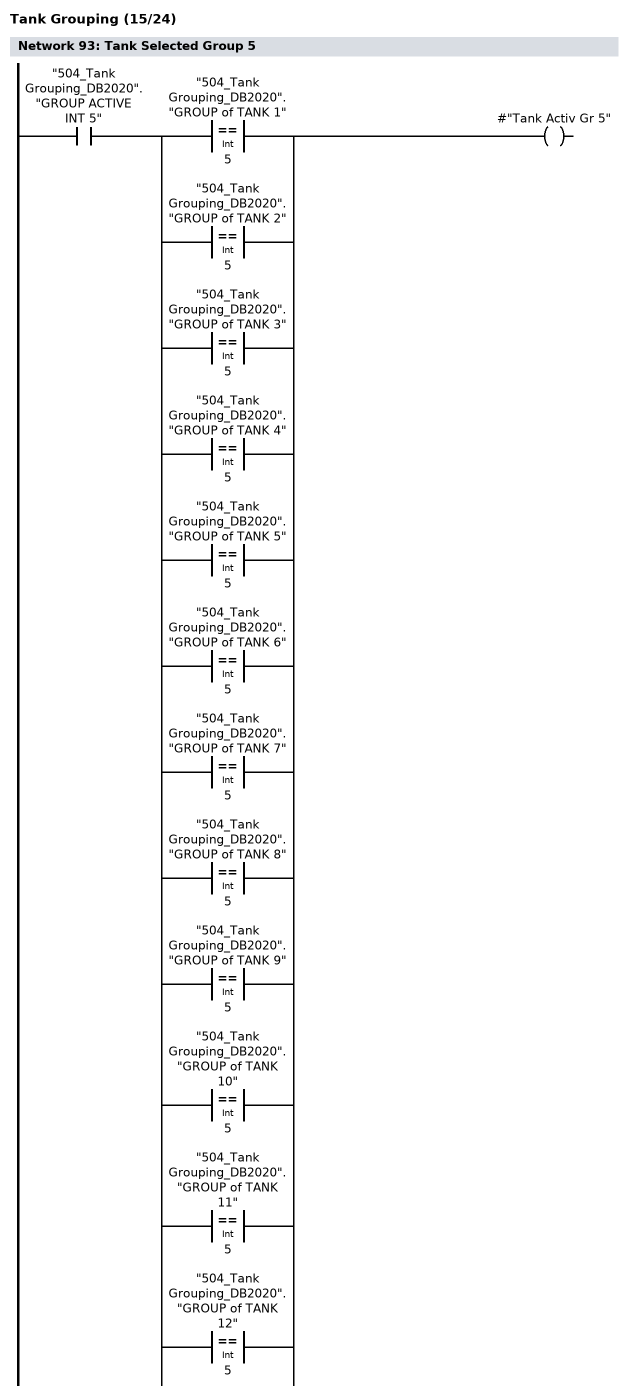
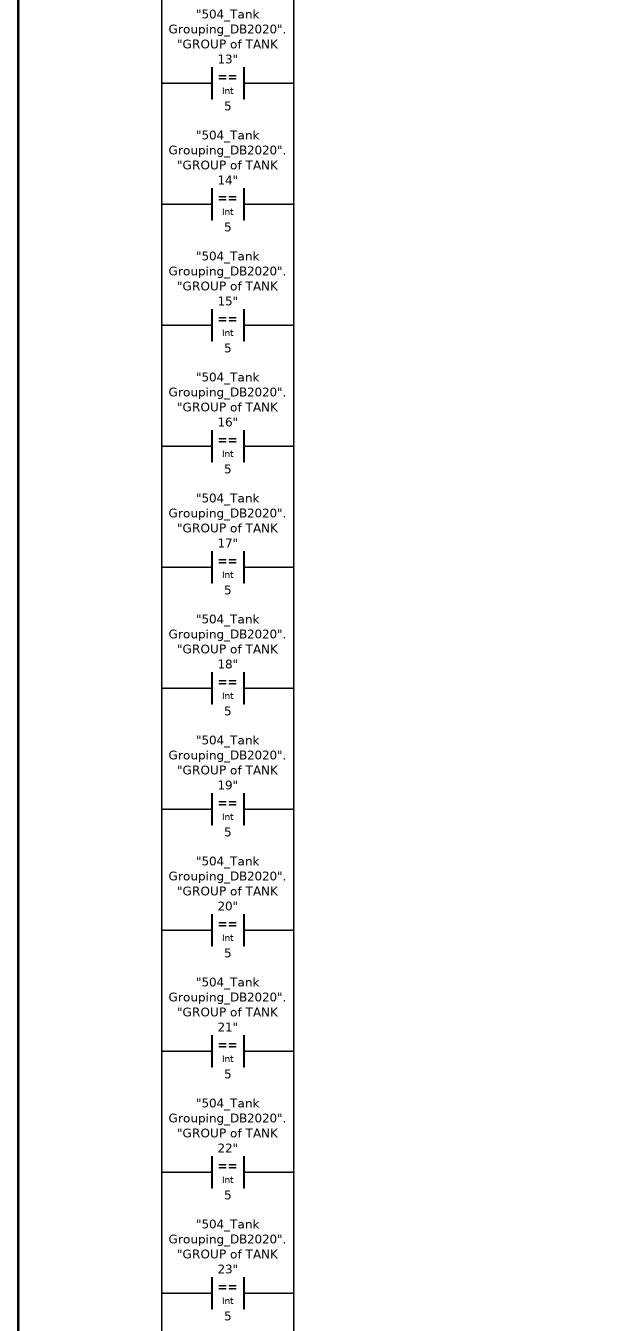
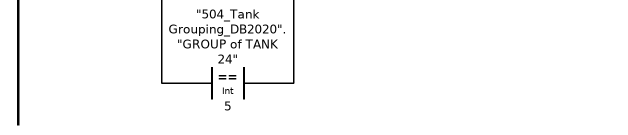
   RUNG wire#powerrail
      Contact( "504_Tank Grouping_DB2020"."GROUP ACTIVE INT 5" )
      wire#w1
      { S7_Templates := "SrcType := Int" } EQ_Contact(in1 := "504_Tank Grouping_DB2020"."GROUP of TANK 1", in2 := 5)
      wire#w2
      Coil( #"Tank Activ Gr 5" )
   END_RUNG
   RUNG wire#w1
      { S7_Templates := "SrcType := Int" } EQ_Contact(in1 := "504_Tank Grouping_DB2020"."GROUP of TANK 2", in2 := 5)
   END_RUNG wire#w2
   RUNG wire#w1
      { S7_Templates := "SrcType := Int" } EQ_Contact(in1 := "504_Tank Grouping_DB2020"."GROUP of TANK 3", in2 := 5)
   END_RUNG wire#w2
   RUNG wire#w1
      { S7_Templates := "SrcType := Int" } EQ_Contact(in1 := "504_Tank Grouping_DB2020"."GROUP of TANK 4", in2 := 5)
   END_RUNG wire#w2
   RUNG wire#w1
      { S7_Templates := "SrcType := Int" } EQ_Contact(in1 := "504_Tank Grouping_DB2020"."GROUP of TANK 5", in2 := 5)
   END_RUNG wire#w2
   RUNG wire#w1
      { S7_Templates := "SrcType := Int" } EQ_Contact(in1 := "504_Tank Grouping_DB2020"."GROUP of TANK 6", in2 := 5)
   END_RUNG wire#w2
   RUNG wire#w1
      { S7_Templates := "SrcType := Int" } EQ_Contact(in1 := "504_Tank Grouping_DB2020"."GROUP of TANK 7", in2 := 5)
   END_RUNG wire#w2
   RUNG wire#w1
      { S7_Templates := "SrcType := Int" } EQ_Contact(in1 := "504_Tank Grouping_DB2020"."GROUP of TANK 8", in2 := 5)
   END_RUNG wire#w2
   RUNG wire#w1
      { S7_Templates := "SrcType := Int" } EQ_Contact(in1 := "504_Tank Grouping_DB2020"."GROUP of TANK 9", in2 := 5)
   END_RUNG wire#w2
   RUNG wire#w1
      { S7_Templates := "SrcType := Int" } EQ_Contact(in1 := "504_Tank Grouping_DB2020"."GROUP of TANK 10", in2 := 5)
   END_RUNG wire#w2
   RUNG wire#w1
      { S7_Templates := "SrcType := Int" } EQ_Contact(in1 := "504_Tank Grouping_DB2020"."GROUP of TANK 11", in2 := 5)
   END_RUNG wire#w2
   RUNG wire#w1
      { S7_Templates := "SrcType := Int" } EQ_Contact(in1 := "504_Tank Grouping_DB2020"."GROUP of TANK 12", in2 := 5)
   END_RUNG wire#w2
   RUNG wire#w1
      { S7_Templates := "SrcType := Int" } EQ_Contact(in1 := "504_Tank Grouping_DB2020"."GROUP of TANK 13", in2 := 5)
   END_RUNG wire#w2
   RUNG wire#w1
      { S7_Templates := "SrcType := Int" } EQ_Contact(in1 := "504_Tank Grouping_DB2020"."GROUP of TANK 14", in2 := 5)
   END_RUNG wire#w2
   RUNG wire#w1
      { S7_Templates := "SrcType := Int" } EQ_Contact(in1 := "504_Tank Grouping_DB2020"."GROUP of TANK 15", in2 := 5)
   END_RUNG wire#w2
   RUNG wire#w1
      { S7_Templates := "SrcType := Int" } EQ_Contact(in1 := "504_Tank Grouping_DB2020"."GROUP of TANK 16", in2 := 5)
   END_RUNG wire#w2
   RUNG wire#w1
      { S7_Templates := "SrcType := Int" } EQ_Contact(in1 := "504_Tank Grouping_DB2020"."GROUP of TANK 17", in2 := 5)
   END_RUNG wire#w2
   RUNG wire#w1
      { S7_Templates := "SrcType := Int" } EQ_Contact(in1 := "504_Tank Grouping_DB2020"."GROUP of TANK 18", in2 := 5)
   END_RUNG wire#w2
   RUNG wire#w1
      { S7_Templates := "SrcType := Int" } EQ_Contact(in1 := "504_Tank Grouping_DB2020"."GROUP of TANK 19", in2 := 5)
   END_RUNG wire#w2
   RUNG wire#w1
      { S7_Templates := "SrcType := Int" } EQ_Contact(in1 := "504_Tank Grouping_DB2020"."GROUP of TANK 20", in2 := 5)
   END_RUNG wire#w2
   RUNG wire#w1
      { S7_Templates := "SrcType := Int" } EQ_Contact(in1 := "504_Tank Grouping_DB2020"."GROUP of TANK 21", in2 := 5)
   END_RUNG wire#w2
   RUNG wire#w1
      { S7_Templates := "SrcType := Int" } EQ_Contact(in1 := "504_Tank Grouping_DB2020"."GROUP of TANK 22", in2 := 5)
   END_RUNG wire#w2
   RUNG wire#w1
      { S7_Templates := "SrcType := Int" } EQ_Contact(in1 := "504_Tank Grouping_DB2020"."GROUP of TANK 23", in2 := 5)
   END_RUNG wire#w2
   RUNG wire#w1
      { S7_Templates := "SrcType := Int" } EQ_Contact(in1 := "504_Tank Grouping_DB2020"."GROUP of TANK 24", in2 := 5)
   END_RUNG wire#w2
   // the same network as SCL:
   #"Tank Activ Gr 5" := "504_Tank Grouping_DB2020"."GROUP ACTIVE INT 5" AND (("504_Tank Grouping_DB2020"."GROUP of TANK 1" = 5) OR ("504_Tank Grouping_DB2020"."GROUP of TANK 2" = 5) OR ("504_Tank Grouping_DB2020"."GROUP of TANK 3" = 5) OR ("504_Tank Grouping_DB2020"."GROUP of TANK 4" = 5) OR ("504_Tank Grouping_DB2020"."GROUP of TANK 5" = 5) OR ("504_Tank Grouping_DB2020"."GROUP of TANK 6" = 5) OR ("504_Tank Grouping_DB2020"."GROUP of TANK 7" = 5) OR ("504_Tank Grouping_DB2020"."GROUP of TANK 8" = 5) OR ("504_Tank Grouping_DB2020"."GROUP of TANK 9" = 5) OR ("504_Tank Grouping_DB2020"."GROUP of TANK 10" = 5) OR ("504_Tank Grouping_DB2020"."GROUP of TANK 11" = 5) OR ("504_Tank Grouping_DB2020"."GROUP of TANK 12" = 5) OR ("504_Tank Grouping_DB2020"."GROUP of TANK 13" = 5) OR ("504_Tank Grouping_DB2020"."GROUP of TANK 14" = 5) OR ("504_Tank Grouping_DB2020"."GROUP of TANK 15" = 5) OR ("504_Tank Grouping_DB2020"."GROUP of TANK 16" = 5) OR ("504_Tank Grouping_DB2020"."GROUP of TANK 17" = 5) OR ("504_Tank Grouping_DB2020"."GROUP of TANK 18" = 5) OR ("504_Tank Grouping_DB2020"."GROUP of TANK 19" = 5) OR ("504_Tank Grouping_DB2020"."GROUP of TANK 20" = 5) OR ("504_Tank Grouping_DB2020"."GROUP of TANK 21" = 5) OR ("504_Tank Grouping_DB2020"."GROUP of TANK 22" = 5) OR ("504_Tank Grouping_DB2020"."GROUP of TANK 23" = 5) OR ("504_Tank Grouping_DB2020"."GROUP of TANK 24" = 5));
END_REGION

REGION Network 94: Tank Selected Group 6
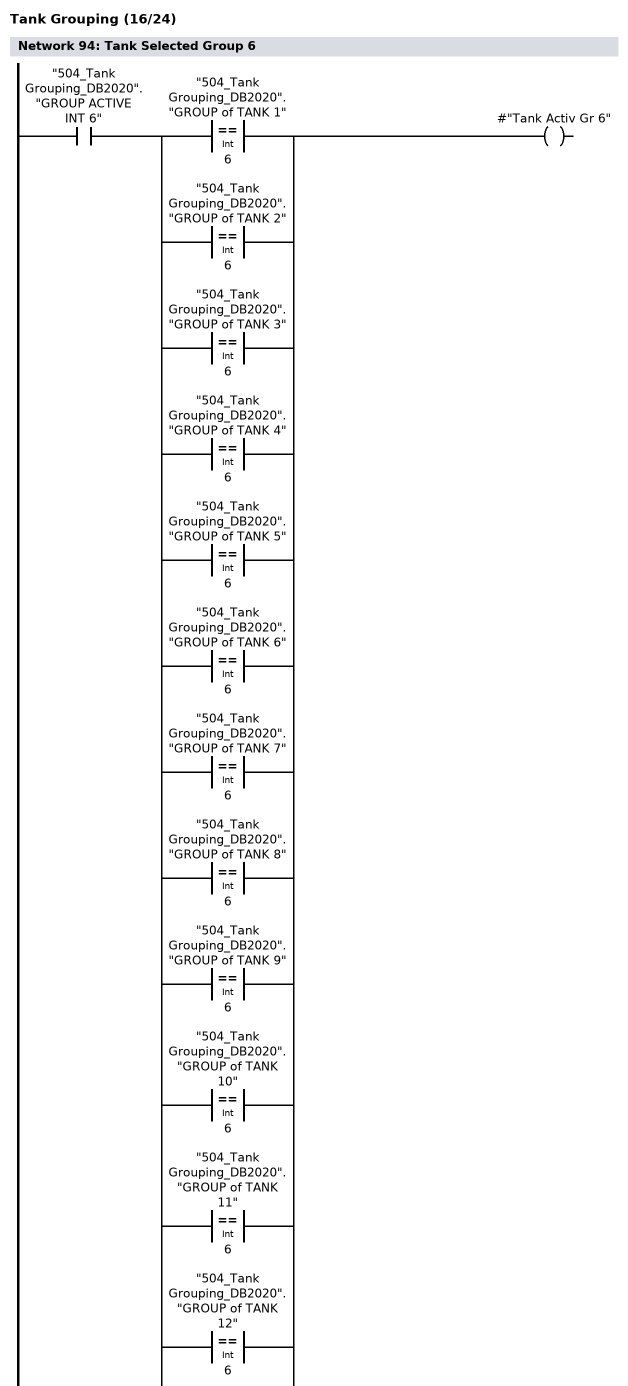
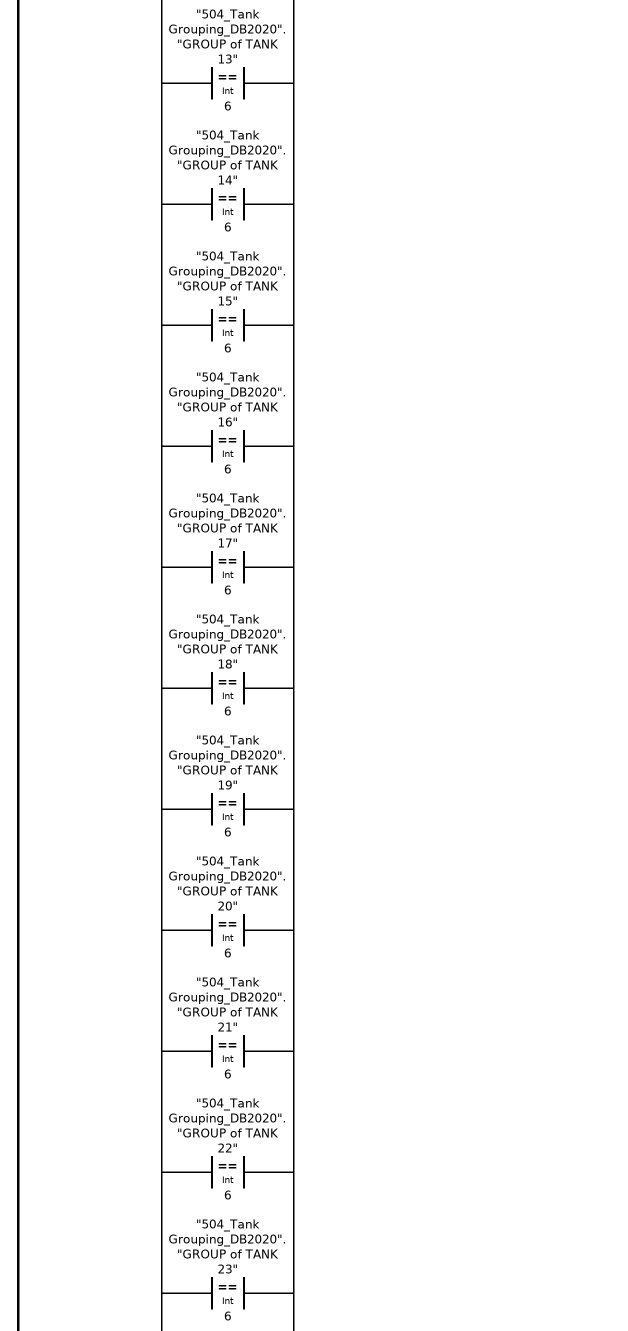
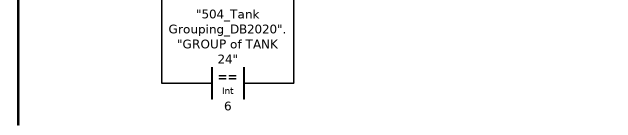
   RUNG wire#powerrail
      Contact( "504_Tank Grouping_DB2020"."GROUP ACTIVE INT 6" )
      wire#w1
      { S7_Templates := "SrcType := Int" } EQ_Contact(in1 := "504_Tank Grouping_DB2020"."GROUP of TANK 1", in2 := 6)
      wire#w2
      Coil( #"Tank Activ Gr 6" )
   END_RUNG
   RUNG wire#w1
      { S7_Templates := "SrcType := Int" } EQ_Contact(in1 := "504_Tank Grouping_DB2020"."GROUP of TANK 2", in2 := 6)
   END_RUNG wire#w2
   RUNG wire#w1
      { S7_Templates := "SrcType := Int" } EQ_Contact(in1 := "504_Tank Grouping_DB2020"."GROUP of TANK 3", in2 := 6)
   END_RUNG wire#w2
   RUNG wire#w1
      { S7_Templates := "SrcType := Int" } EQ_Contact(in1 := "504_Tank Grouping_DB2020"."GROUP of TANK 4", in2 := 6)
   END_RUNG wire#w2
   RUNG wire#w1
      { S7_Templates := "SrcType := Int" } EQ_Contact(in1 := "504_Tank Grouping_DB2020"."GROUP of TANK 5", in2 := 6)
   END_RUNG wire#w2
   RUNG wire#w1
      { S7_Templates := "SrcType := Int" } EQ_Contact(in1 := "504_Tank Grouping_DB2020"."GROUP of TANK 6", in2 := 6)
   END_RUNG wire#w2
   RUNG wire#w1
      { S7_Templates := "SrcType := Int" } EQ_Contact(in1 := "504_Tank Grouping_DB2020"."GROUP of TANK 7", in2 := 6)
   END_RUNG wire#w2
   RUNG wire#w1
      { S7_Templates := "SrcType := Int" } EQ_Contact(in1 := "504_Tank Grouping_DB2020"."GROUP of TANK 8", in2 := 6)
   END_RUNG wire#w2
   RUNG wire#w1
      { S7_Templates := "SrcType := Int" } EQ_Contact(in1 := "504_Tank Grouping_DB2020"."GROUP of TANK 9", in2 := 6)
   END_RUNG wire#w2
   RUNG wire#w1
      { S7_Templates := "SrcType := Int" } EQ_Contact(in1 := "504_Tank Grouping_DB2020"."GROUP of TANK 10", in2 := 6)
   END_RUNG wire#w2
   RUNG wire#w1
      { S7_Templates := "SrcType := Int" } EQ_Contact(in1 := "504_Tank Grouping_DB2020"."GROUP of TANK 11", in2 := 6)
   END_RUNG wire#w2
   RUNG wire#w1
      { S7_Templates := "SrcType := Int" } EQ_Contact(in1 := "504_Tank Grouping_DB2020"."GROUP of TANK 12", in2 := 6)
   END_RUNG wire#w2
   RUNG wire#w1
      { S7_Templates := "SrcType := Int" } EQ_Contact(in1 := "504_Tank Grouping_DB2020"."GROUP of TANK 13", in2 := 6)
   END_RUNG wire#w2
   RUNG wire#w1
      { S7_Templates := "SrcType := Int" } EQ_Contact(in1 := "504_Tank Grouping_DB2020"."GROUP of TANK 14", in2 := 6)
   END_RUNG wire#w2
   RUNG wire#w1
      { S7_Templates := "SrcType := Int" } EQ_Contact(in1 := "504_Tank Grouping_DB2020"."GROUP of TANK 15", in2 := 6)
   END_RUNG wire#w2
   RUNG wire#w1
      { S7_Templates := "SrcType := Int" } EQ_Contact(in1 := "504_Tank Grouping_DB2020"."GROUP of TANK 16", in2 := 6)
   END_RUNG wire#w2
   RUNG wire#w1
      { S7_Templates := "SrcType := Int" } EQ_Contact(in1 := "504_Tank Grouping_DB2020"."GROUP of TANK 17", in2 := 6)
   END_RUNG wire#w2
   RUNG wire#w1
      { S7_Templates := "SrcType := Int" } EQ_Contact(in1 := "504_Tank Grouping_DB2020"."GROUP of TANK 18", in2 := 6)
   END_RUNG wire#w2
   RUNG wire#w1
      { S7_Templates := "SrcType := Int" } EQ_Contact(in1 := "504_Tank Grouping_DB2020"."GROUP of TANK 19", in2 := 6)
   END_RUNG wire#w2
   RUNG wire#w1
      { S7_Templates := "SrcType := Int" } EQ_Contact(in1 := "504_Tank Grouping_DB2020"."GROUP of TANK 20", in2 := 6)
   END_RUNG wire#w2
   RUNG wire#w1
      { S7_Templates := "SrcType := Int" } EQ_Contact(in1 := "504_Tank Grouping_DB2020"."GROUP of TANK 21", in2 := 6)
   END_RUNG wire#w2
   RUNG wire#w1
      { S7_Templates := "SrcType := Int" } EQ_Contact(in1 := "504_Tank Grouping_DB2020"."GROUP of TANK 22", in2 := 6)
   END_RUNG wire#w2
   RUNG wire#w1
      { S7_Templates := "SrcType := Int" } EQ_Contact(in1 := "504_Tank Grouping_DB2020"."GROUP of TANK 23", in2 := 6)
   END_RUNG wire#w2
   RUNG wire#w1
      { S7_Templates := "SrcType := Int" } EQ_Contact(in1 := "504_Tank Grouping_DB2020"."GROUP of TANK 24", in2 := 6)
   END_RUNG wire#w2
   // the same network as SCL:
   #"Tank Activ Gr 6" := "504_Tank Grouping_DB2020"."GROUP ACTIVE INT 6" AND (("504_Tank Grouping_DB2020"."GROUP of TANK 1" = 6) OR ("504_Tank Grouping_DB2020"."GROUP of TANK 2" = 6) OR ("504_Tank Grouping_DB2020"."GROUP of TANK 3" = 6) OR ("504_Tank Grouping_DB2020"."GROUP of TANK 4" = 6) OR ("504_Tank Grouping_DB2020"."GROUP of TANK 5" = 6) OR ("504_Tank Grouping_DB2020"."GROUP of TANK 6" = 6) OR ("504_Tank Grouping_DB2020"."GROUP of TANK 7" = 6) OR ("504_Tank Grouping_DB2020"."GROUP of TANK 8" = 6) OR ("504_Tank Grouping_DB2020"."GROUP of TANK 9" = 6) OR ("504_Tank Grouping_DB2020"."GROUP of TANK 10" = 6) OR ("504_Tank Grouping_DB2020"."GROUP of TANK 11" = 6) OR ("504_Tank Grouping_DB2020"."GROUP of TANK 12" = 6) OR ("504_Tank Grouping_DB2020"."GROUP of TANK 13" = 6) OR ("504_Tank Grouping_DB2020"."GROUP of TANK 14" = 6) OR ("504_Tank Grouping_DB2020"."GROUP of TANK 15" = 6) OR ("504_Tank Grouping_DB2020"."GROUP of TANK 16" = 6) OR ("504_Tank Grouping_DB2020"."GROUP of TANK 17" = 6) OR ("504_Tank Grouping_DB2020"."GROUP of TANK 18" = 6) OR ("504_Tank Grouping_DB2020"."GROUP of TANK 19" = 6) OR ("504_Tank Grouping_DB2020"."GROUP of TANK 20" = 6) OR ("504_Tank Grouping_DB2020"."GROUP of TANK 21" = 6) OR ("504_Tank Grouping_DB2020"."GROUP of TANK 22" = 6) OR ("504_Tank Grouping_DB2020"."GROUP of TANK 23" = 6) OR ("504_Tank Grouping_DB2020"."GROUP of TANK 24" = 6));
END_REGION

REGION Network 95: Tank Selected Group 7
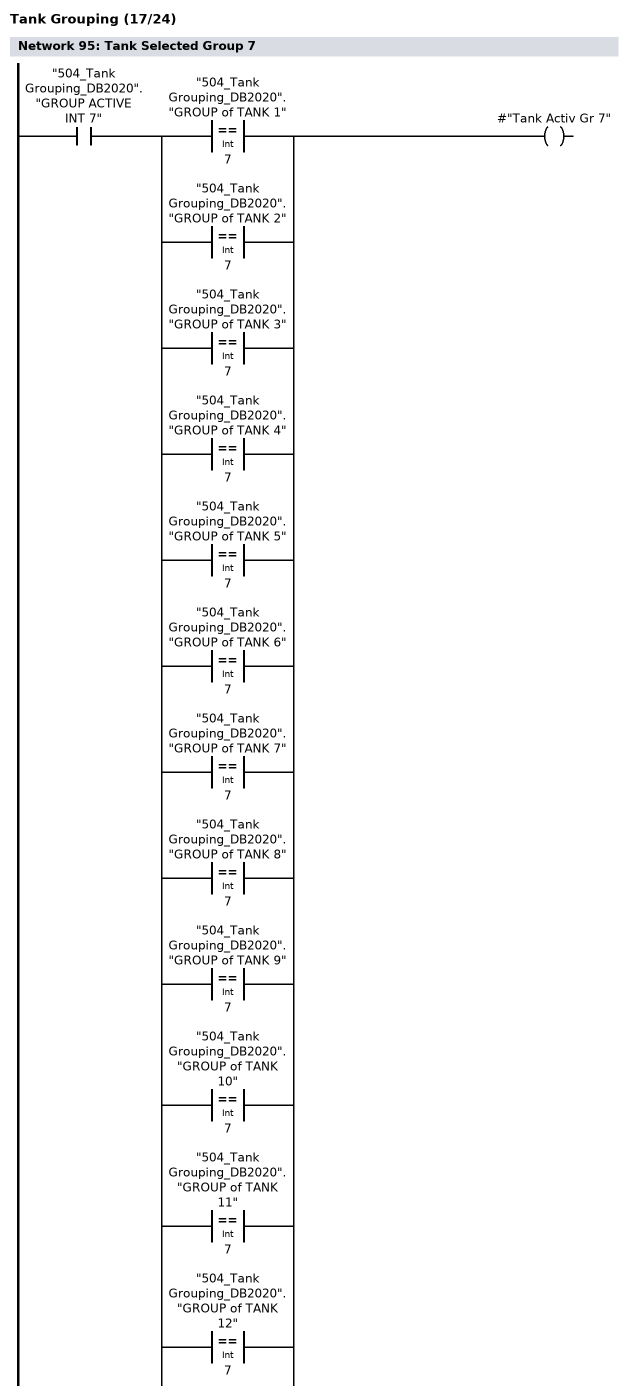
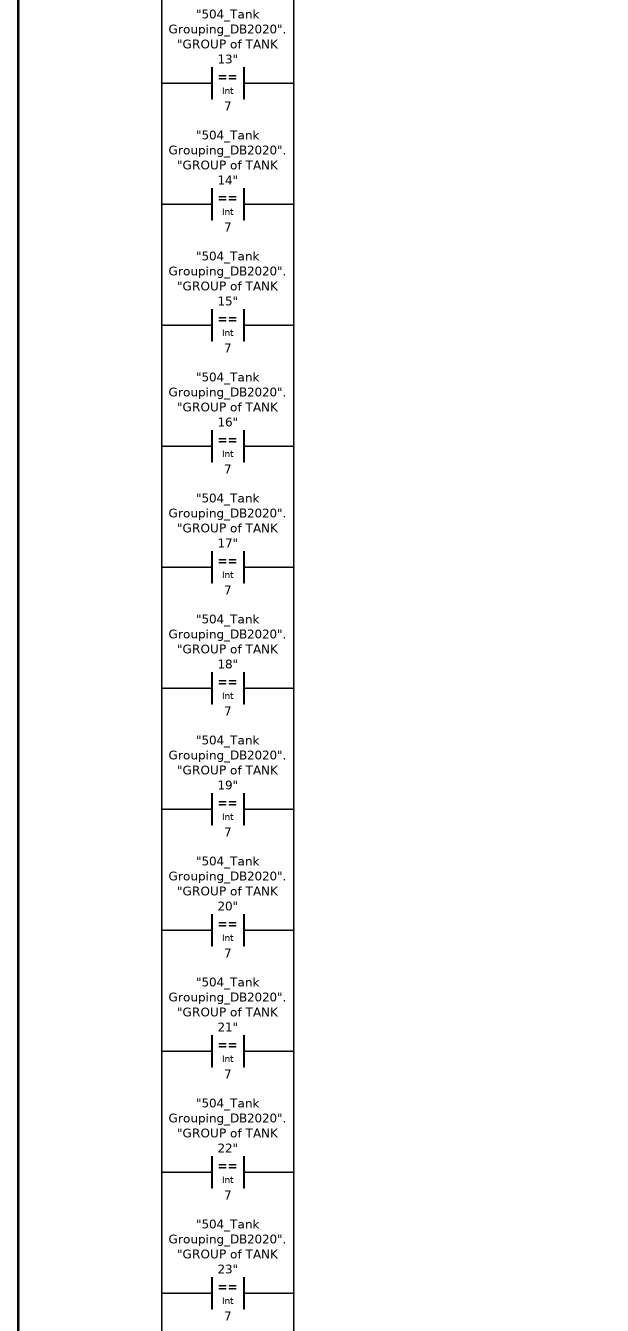
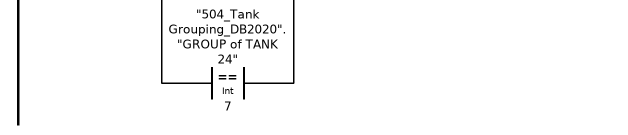
   RUNG wire#powerrail
      Contact( "504_Tank Grouping_DB2020"."GROUP ACTIVE INT 7" )
      wire#w1
      { S7_Templates := "SrcType := Int" } EQ_Contact(in1 := "504_Tank Grouping_DB2020"."GROUP of TANK 1", in2 := 7)
      wire#w2
      Coil( #"Tank Activ Gr 7" )
   END_RUNG
   RUNG wire#w1
      { S7_Templates := "SrcType := Int" } EQ_Contact(in1 := "504_Tank Grouping_DB2020"."GROUP of TANK 2", in2 := 7)
   END_RUNG wire#w2
   RUNG wire#w1
      { S7_Templates := "SrcType := Int" } EQ_Contact(in1 := "504_Tank Grouping_DB2020"."GROUP of TANK 3", in2 := 7)
   END_RUNG wire#w2
   RUNG wire#w1
      { S7_Templates := "SrcType := Int" } EQ_Contact(in1 := "504_Tank Grouping_DB2020"."GROUP of TANK 4", in2 := 7)
   END_RUNG wire#w2
   RUNG wire#w1
      { S7_Templates := "SrcType := Int" } EQ_Contact(in1 := "504_Tank Grouping_DB2020"."GROUP of TANK 5", in2 := 7)
   END_RUNG wire#w2
   RUNG wire#w1
      { S7_Templates := "SrcType := Int" } EQ_Contact(in1 := "504_Tank Grouping_DB2020"."GROUP of TANK 6", in2 := 7)
   END_RUNG wire#w2
   RUNG wire#w1
      { S7_Templates := "SrcType := Int" } EQ_Contact(in1 := "504_Tank Grouping_DB2020"."GROUP of TANK 7", in2 := 7)
   END_RUNG wire#w2
   RUNG wire#w1
      { S7_Templates := "SrcType := Int" } EQ_Contact(in1 := "504_Tank Grouping_DB2020"."GROUP of TANK 8", in2 := 7)
   END_RUNG wire#w2
   RUNG wire#w1
      { S7_Templates := "SrcType := Int" } EQ_Contact(in1 := "504_Tank Grouping_DB2020"."GROUP of TANK 9", in2 := 7)
   END_RUNG wire#w2
   RUNG wire#w1
      { S7_Templates := "SrcType := Int" } EQ_Contact(in1 := "504_Tank Grouping_DB2020"."GROUP of TANK 10", in2 := 7)
   END_RUNG wire#w2
   RUNG wire#w1
      { S7_Templates := "SrcType := Int" } EQ_Contact(in1 := "504_Tank Grouping_DB2020"."GROUP of TANK 11", in2 := 7)
   END_RUNG wire#w2
   RUNG wire#w1
      { S7_Templates := "SrcType := Int" } EQ_Contact(in1 := "504_Tank Grouping_DB2020"."GROUP of TANK 12", in2 := 7)
   END_RUNG wire#w2
   RUNG wire#w1
      { S7_Templates := "SrcType := Int" } EQ_Contact(in1 := "504_Tank Grouping_DB2020"."GROUP of TANK 13", in2 := 7)
   END_RUNG wire#w2
   RUNG wire#w1
      { S7_Templates := "SrcType := Int" } EQ_Contact(in1 := "504_Tank Grouping_DB2020"."GROUP of TANK 14", in2 := 7)
   END_RUNG wire#w2
   RUNG wire#w1
      { S7_Templates := "SrcType := Int" } EQ_Contact(in1 := "504_Tank Grouping_DB2020"."GROUP of TANK 15", in2 := 7)
   END_RUNG wire#w2
   RUNG wire#w1
      { S7_Templates := "SrcType := Int" } EQ_Contact(in1 := "504_Tank Grouping_DB2020"."GROUP of TANK 16", in2 := 7)
   END_RUNG wire#w2
   RUNG wire#w1
      { S7_Templates := "SrcType := Int" } EQ_Contact(in1 := "504_Tank Grouping_DB2020"."GROUP of TANK 17", in2 := 7)
   END_RUNG wire#w2
   RUNG wire#w1
      { S7_Templates := "SrcType := Int" } EQ_Contact(in1 := "504_Tank Grouping_DB2020"."GROUP of TANK 18", in2 := 7)
   END_RUNG wire#w2
   RUNG wire#w1
      { S7_Templates := "SrcType := Int" } EQ_Contact(in1 := "504_Tank Grouping_DB2020"."GROUP of TANK 19", in2 := 7)
   END_RUNG wire#w2
   RUNG wire#w1
      { S7_Templates := "SrcType := Int" } EQ_Contact(in1 := "504_Tank Grouping_DB2020"."GROUP of TANK 20", in2 := 7)
   END_RUNG wire#w2
   RUNG wire#w1
      { S7_Templates := "SrcType := Int" } EQ_Contact(in1 := "504_Tank Grouping_DB2020"."GROUP of TANK 21", in2 := 7)
   END_RUNG wire#w2
   RUNG wire#w1
      { S7_Templates := "SrcType := Int" } EQ_Contact(in1 := "504_Tank Grouping_DB2020"."GROUP of TANK 22", in2 := 7)
   END_RUNG wire#w2
   RUNG wire#w1
      { S7_Templates := "SrcType := Int" } EQ_Contact(in1 := "504_Tank Grouping_DB2020"."GROUP of TANK 23", in2 := 7)
   END_RUNG wire#w2
   RUNG wire#w1
      { S7_Templates := "SrcType := Int" } EQ_Contact(in1 := "504_Tank Grouping_DB2020"."GROUP of TANK 24", in2 := 7)
   END_RUNG wire#w2
   // the same network as SCL:
   #"Tank Activ Gr 7" := "504_Tank Grouping_DB2020"."GROUP ACTIVE INT 7" AND (("504_Tank Grouping_DB2020"."GROUP of TANK 1" = 7) OR ("504_Tank Grouping_DB2020"."GROUP of TANK 2" = 7) OR ("504_Tank Grouping_DB2020"."GROUP of TANK 3" = 7) OR ("504_Tank Grouping_DB2020"."GROUP of TANK 4" = 7) OR ("504_Tank Grouping_DB2020"."GROUP of TANK 5" = 7) OR ("504_Tank Grouping_DB2020"."GROUP of TANK 6" = 7) OR ("504_Tank Grouping_DB2020"."GROUP of TANK 7" = 7) OR ("504_Tank Grouping_DB2020"."GROUP of TANK 8" = 7) OR ("504_Tank Grouping_DB2020"."GROUP of TANK 9" = 7) OR ("504_Tank Grouping_DB2020"."GROUP of TANK 10" = 7) OR ("504_Tank Grouping_DB2020"."GROUP of TANK 11" = 7) OR ("504_Tank Grouping_DB2020"."GROUP of TANK 12" = 7) OR ("504_Tank Grouping_DB2020"."GROUP of TANK 13" = 7) OR ("504_Tank Grouping_DB2020"."GROUP of TANK 14" = 7) OR ("504_Tank Grouping_DB2020"."GROUP of TANK 15" = 7) OR ("504_Tank Grouping_DB2020"."GROUP of TANK 16" = 7) OR ("504_Tank Grouping_DB2020"."GROUP of TANK 17" = 7) OR ("504_Tank Grouping_DB2020"."GROUP of TANK 18" = 7) OR ("504_Tank Grouping_DB2020"."GROUP of TANK 19" = 7) OR ("504_Tank Grouping_DB2020"."GROUP of TANK 20" = 7) OR ("504_Tank Grouping_DB2020"."GROUP of TANK 21" = 7) OR ("504_Tank Grouping_DB2020"."GROUP of TANK 22" = 7) OR ("504_Tank Grouping_DB2020"."GROUP of TANK 23" = 7) OR ("504_Tank Grouping_DB2020"."GROUP of TANK 24" = 7));
END_REGION

REGION Network 96: Tank Selected Group 8
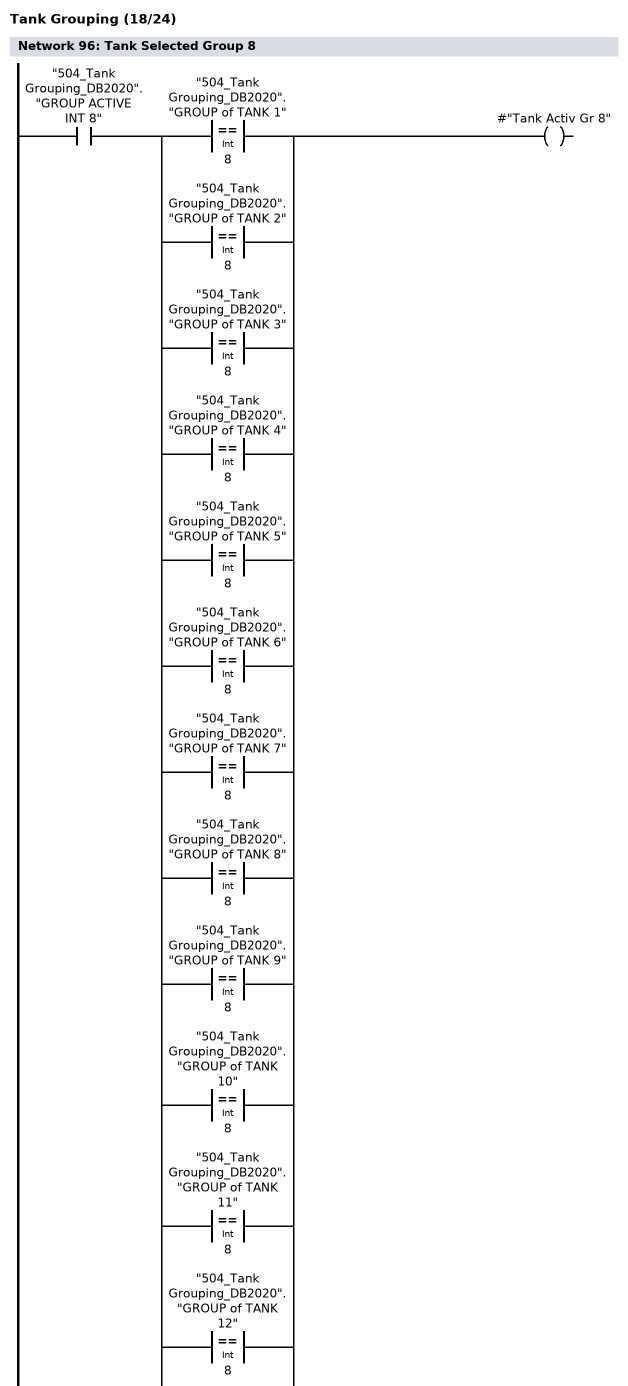
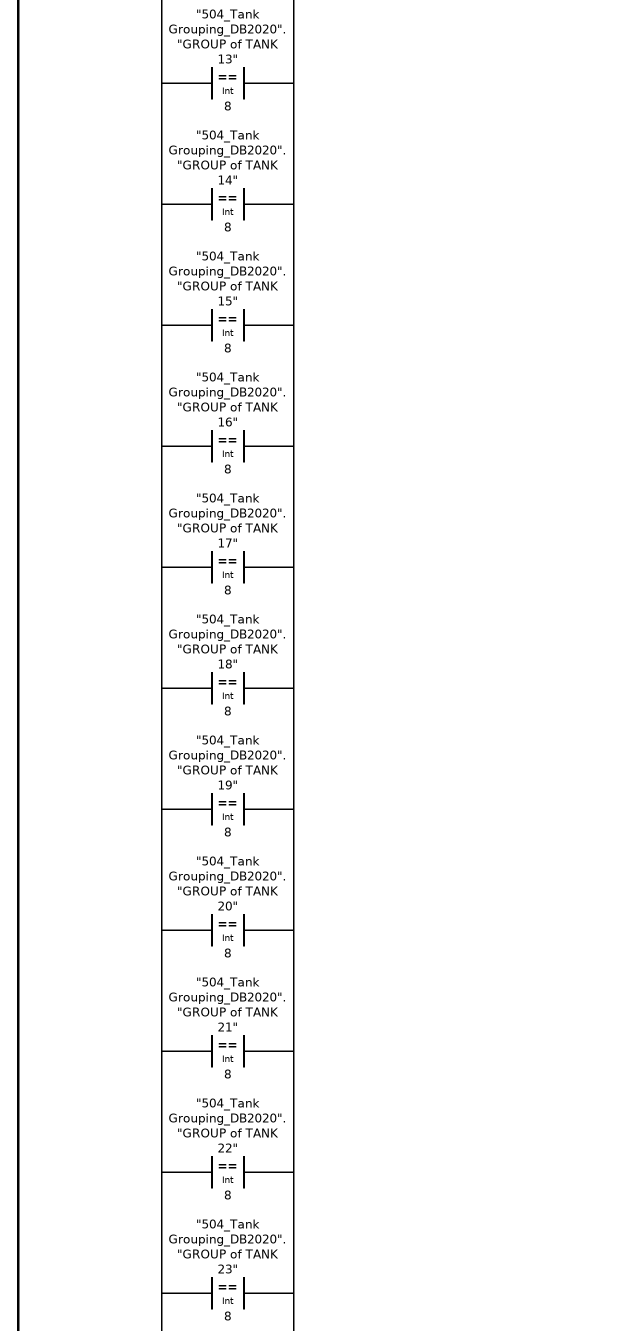
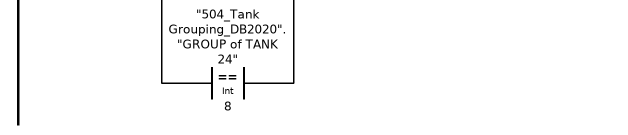
   RUNG wire#powerrail
      Contact( "504_Tank Grouping_DB2020"."GROUP ACTIVE INT 8" )
      wire#w1
      { S7_Templates := "SrcType := Int" } EQ_Contact(in1 := "504_Tank Grouping_DB2020"."GROUP of TANK 1", in2 := 8)
      wire#w2
      Coil( #"Tank Activ Gr 8" )
   END_RUNG
   RUNG wire#w1
      { S7_Templates := "SrcType := Int" } EQ_Contact(in1 := "504_Tank Grouping_DB2020"."GROUP of TANK 2", in2 := 8)
   END_RUNG wire#w2
   RUNG wire#w1
      { S7_Templates := "SrcType := Int" } EQ_Contact(in1 := "504_Tank Grouping_DB2020"."GROUP of TANK 3", in2 := 8)
   END_RUNG wire#w2
   RUNG wire#w1
      { S7_Templates := "SrcType := Int" } EQ_Contact(in1 := "504_Tank Grouping_DB2020"."GROUP of TANK 4", in2 := 8)
   END_RUNG wire#w2
   RUNG wire#w1
      { S7_Templates := "SrcType := Int" } EQ_Contact(in1 := "504_Tank Grouping_DB2020"."GROUP of TANK 5", in2 := 8)
   END_RUNG wire#w2
   RUNG wire#w1
      { S7_Templates := "SrcType := Int" } EQ_Contact(in1 := "504_Tank Grouping_DB2020"."GROUP of TANK 6", in2 := 8)
   END_RUNG wire#w2
   RUNG wire#w1
      { S7_Templates := "SrcType := Int" } EQ_Contact(in1 := "504_Tank Grouping_DB2020"."GROUP of TANK 7", in2 := 8)
   END_RUNG wire#w2
   RUNG wire#w1
      { S7_Templates := "SrcType := Int" } EQ_Contact(in1 := "504_Tank Grouping_DB2020"."GROUP of TANK 8", in2 := 8)
   END_RUNG wire#w2
   RUNG wire#w1
      { S7_Templates := "SrcType := Int" } EQ_Contact(in1 := "504_Tank Grouping_DB2020"."GROUP of TANK 9", in2 := 8)
   END_RUNG wire#w2
   RUNG wire#w1
      { S7_Templates := "SrcType := Int" } EQ_Contact(in1 := "504_Tank Grouping_DB2020"."GROUP of TANK 10", in2 := 8)
   END_RUNG wire#w2
   RUNG wire#w1
      { S7_Templates := "SrcType := Int" } EQ_Contact(in1 := "504_Tank Grouping_DB2020"."GROUP of TANK 11", in2 := 8)
   END_RUNG wire#w2
   RUNG wire#w1
      { S7_Templates := "SrcType := Int" } EQ_Contact(in1 := "504_Tank Grouping_DB2020"."GROUP of TANK 12", in2 := 8)
   END_RUNG wire#w2
   RUNG wire#w1
      { S7_Templates := "SrcType := Int" } EQ_Contact(in1 := "504_Tank Grouping_DB2020"."GROUP of TANK 13", in2 := 8)
   END_RUNG wire#w2
   RUNG wire#w1
      { S7_Templates := "SrcType := Int" } EQ_Contact(in1 := "504_Tank Grouping_DB2020"."GROUP of TANK 14", in2 := 8)
   END_RUNG wire#w2
   RUNG wire#w1
      { S7_Templates := "SrcType := Int" } EQ_Contact(in1 := "504_Tank Grouping_DB2020"."GROUP of TANK 15", in2 := 8)
   END_RUNG wire#w2
   RUNG wire#w1
      { S7_Templates := "SrcType := Int" } EQ_Contact(in1 := "504_Tank Grouping_DB2020"."GROUP of TANK 16", in2 := 8)
   END_RUNG wire#w2
   RUNG wire#w1
      { S7_Templates := "SrcType := Int" } EQ_Contact(in1 := "504_Tank Grouping_DB2020"."GROUP of TANK 17", in2 := 8)
   END_RUNG wire#w2
   RUNG wire#w1
      { S7_Templates := "SrcType := Int" } EQ_Contact(in1 := "504_Tank Grouping_DB2020"."GROUP of TANK 18", in2 := 8)
   END_RUNG wire#w2
   RUNG wire#w1
      { S7_Templates := "SrcType := Int" } EQ_Contact(in1 := "504_Tank Grouping_DB2020"."GROUP of TANK 19", in2 := 8)
   END_RUNG wire#w2
   RUNG wire#w1
      { S7_Templates := "SrcType := Int" } EQ_Contact(in1 := "504_Tank Grouping_DB2020"."GROUP of TANK 20", in2 := 8)
   END_RUNG wire#w2
   RUNG wire#w1
      { S7_Templates := "SrcType := Int" } EQ_Contact(in1 := "504_Tank Grouping_DB2020"."GROUP of TANK 21", in2 := 8)
   END_RUNG wire#w2
   RUNG wire#w1
      { S7_Templates := "SrcType := Int" } EQ_Contact(in1 := "504_Tank Grouping_DB2020"."GROUP of TANK 22", in2 := 8)
   END_RUNG wire#w2
   RUNG wire#w1
      { S7_Templates := "SrcType := Int" } EQ_Contact(in1 := "504_Tank Grouping_DB2020"."GROUP of TANK 23", in2 := 8)
   END_RUNG wire#w2
   RUNG wire#w1
      { S7_Templates := "SrcType := Int" } EQ_Contact(in1 := "504_Tank Grouping_DB2020"."GROUP of TANK 24", in2 := 8)
   END_RUNG wire#w2
   // the same network as SCL:
   #"Tank Activ Gr 8" := "504_Tank Grouping_DB2020"."GROUP ACTIVE INT 8" AND (("504_Tank Grouping_DB2020"."GROUP of TANK 1" = 8) OR ("504_Tank Grouping_DB2020"."GROUP of TANK 2" = 8) OR ("504_Tank Grouping_DB2020"."GROUP of TANK 3" = 8) OR ("504_Tank Grouping_DB2020"."GROUP of TANK 4" = 8) OR ("504_Tank Grouping_DB2020"."GROUP of TANK 5" = 8) OR ("504_Tank Grouping_DB2020"."GROUP of TANK 6" = 8) OR ("504_Tank Grouping_DB2020"."GROUP of TANK 7" = 8) OR ("504_Tank Grouping_DB2020"."GROUP of TANK 8" = 8) OR ("504_Tank Grouping_DB2020"."GROUP of TANK 9" = 8) OR ("504_Tank Grouping_DB2020"."GROUP of TANK 10" = 8) OR ("504_Tank Grouping_DB2020"."GROUP of TANK 11" = 8) OR ("504_Tank Grouping_DB2020"."GROUP of TANK 12" = 8) OR ("504_Tank Grouping_DB2020"."GROUP of TANK 13" = 8) OR ("504_Tank Grouping_DB2020"."GROUP of TANK 14" = 8) OR ("504_Tank Grouping_DB2020"."GROUP of TANK 15" = 8) OR ("504_Tank Grouping_DB2020"."GROUP of TANK 16" = 8) OR ("504_Tank Grouping_DB2020"."GROUP of TANK 17" = 8) OR ("504_Tank Grouping_DB2020"."GROUP of TANK 18" = 8) OR ("504_Tank Grouping_DB2020"."GROUP of TANK 19" = 8) OR ("504_Tank Grouping_DB2020"."GROUP of TANK 20" = 8) OR ("504_Tank Grouping_DB2020"."GROUP of TANK 21" = 8) OR ("504_Tank Grouping_DB2020"."GROUP of TANK 22" = 8) OR ("504_Tank Grouping_DB2020"."GROUP of TANK 23" = 8) OR ("504_Tank Grouping_DB2020"."GROUP of TANK 24" = 8));
END_REGION

REGION Network 97: Tank Selected Group 9